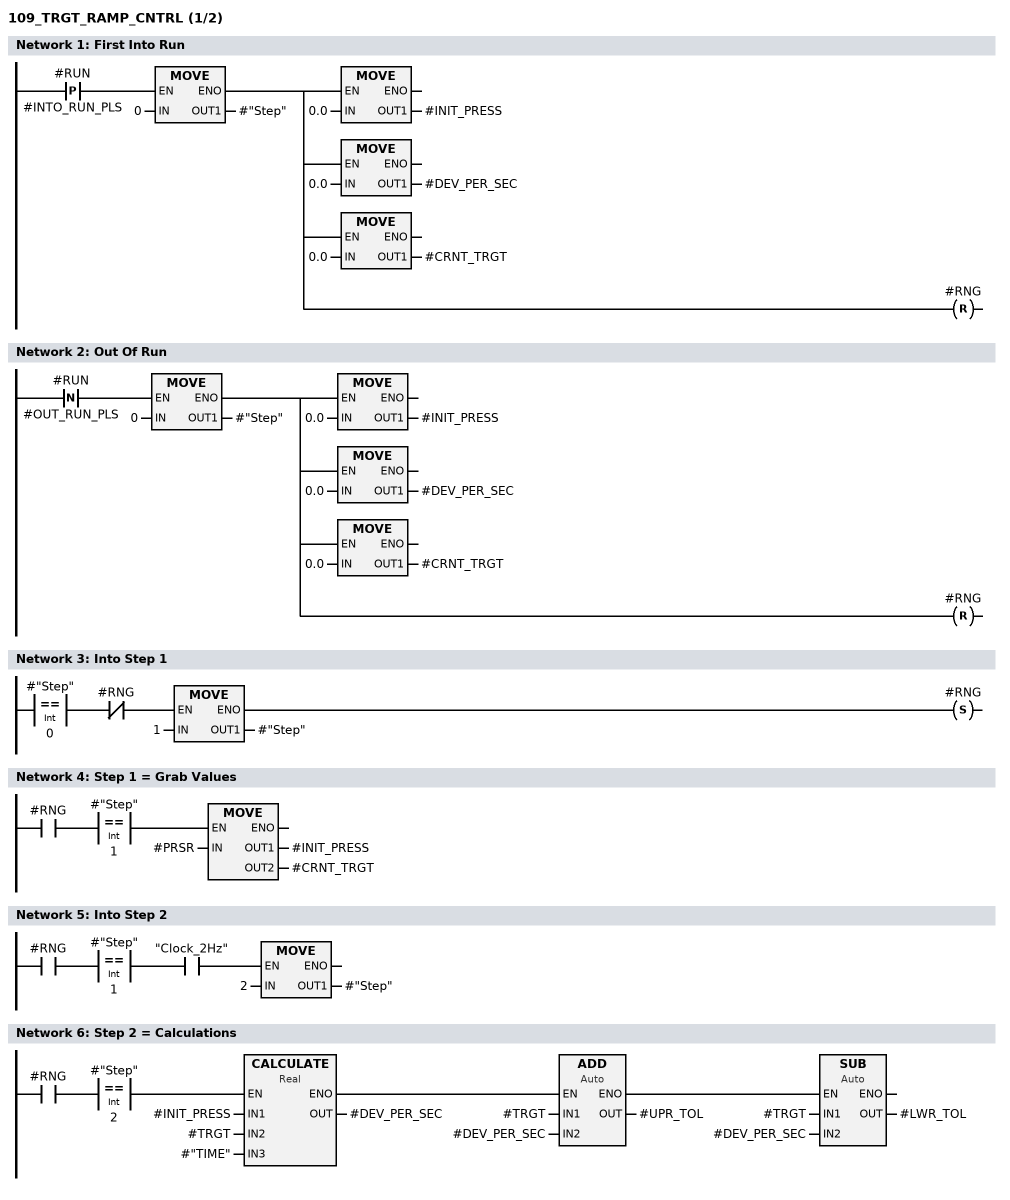
   RUNG wire#powerrail
      P_Contact(operand := #RUN, bit := #INTO_RUN_PLS)
      Move(in := 0, out1 => #"Step")
      wire#w1
      Move(in := 0.0, out1 => #INIT_PRESS)
   END_RUNG
   RUNG wire#w1
      Move(in := 0.0, out1 => #DEV_PER_SEC)
   END_RUNG
   RUNG wire#w1
      Move(in := 0.0, out1 => #CRNT_TRGT)
   END_RUNG
   RUNG wire#w1
      R_Coil( #RNG )
   END_RUNG
   // the same network as SCL:
   #_w1 := #RUN AND NOT #INTO_RUN_PLS;   // rising edge of #RUN
   #INTO_RUN_PLS := #RUN;
   IF #_w1 THEN
       #"Step" := 0;
       #INIT_PRESS := 0.0;
       #DEV_PER_SEC := 0.0;
       #CRNT_TRGT := 0.0;
       #RNG := FALSE;
   END_IF;
END_REGION

REGION Network 2: Out Of Run
   RUNG wire#powerrail
      N_Contact(operand := #RUN, bit := #OUT_RUN_PLS)
      Move(in := 0, out1 => #"Step")
      wire#w1
      Move(in := 0.0, out1 => #INIT_PRESS)
   END_RUNG
   RUNG wire#w1
      Move(in := 0.0, out1 => #DEV_PER_SEC)
   END_RUNG
   RUNG wire#w1
      Move(in := 0.0, out1 => #CRNT_TRGT)
   END_RUNG
   RUNG wire#w1
      R_Coil( #RNG )
   END_RUNG
   // the same network as SCL:
   #_w1 := NOT #RUN AND #OUT_RUN_PLS;   // falling edge of #RUN
   #OUT_RUN_PLS := #RUN;
   IF #_w1 THEN
       #"Step" := 0;
       #INIT_PRESS := 0.0;
       #DEV_PER_SEC := 0.0;
       #CRNT_TRGT := 0.0;
       #RNG := FALSE;
   END_IF;
END_REGION

REGION Network 3: Into Step 1
   RUNG wire#powerrail
      { S7_Templates := "SrcType := Int" } EQ_Contact(in1 := #"Step", in2 := 0)
      I_Contact( #RNG )
      Move(in := 1, out1 => #"Step")
      S_Coil( #RNG )
   END_RUNG
   // the same network as SCL:
   #_w1 := (#"Step" = 0) AND NOT #RNG;
   IF #_w1 THEN
       #"Step" := 1;
       #RNG := TRUE;
   END_IF;
END_REGION

REGION Network 4: Step 1 = Grab Values
   RUNG wire#powerrail
      Contact( #RNG )
      { S7_Templates := "SrcType := Int" } EQ_Contact(in1 := #"Step", in2 := 1)
      Move(in := #PRSR, out1 => #INIT_PRESS, out2 => #CRNT_TRGT)
   END_RUNG
   // the same network as SCL:
   IF #RNG AND (#"Step" = 1) THEN
       #INIT_PRESS := #PRSR;
       #CRNT_TRGT := #PRSR;
   END_IF;
END_REGION

REGION Network 5: Into Step 2
   RUNG wire#powerrail
      Contact( #RNG )
      { S7_Templates := "SrcType := Int" } EQ_Contact(in1 := #"Step", in2 := 1)
      Contact( "Clock_2Hz" )
      Move(in := 2, out1 => #"Step")
   END_RUNG
   // the same network as SCL:
   IF #RNG AND (#"Step" = 1) AND "Clock_2Hz" THEN #"Step" := 2; END_IF;
END_REGION

REGION Network 6: Step 2 = Calculations
   RUNG wire#powerrail
      Contact( #RNG )
      { S7_Templates := "SrcType := Int" } EQ_Contact(in1 := #"Step", in2 := 2)
      { S7_Templates := "SrcType := Real"; S7_Expression := "(IN2-IN1)/IN3" } Calculate(in1 := #INIT_PRESS, in2 := #TRGT, in3 := #"TIME", out => #DEV_PER_SEC)
      Add(in1 := #TRGT, in2 := #DEV_PER_SEC, out => #UPR_TOL)
      Sub(in1 := #TRGT, in2 := #DEV_PER_SEC, out => #LWR_TOL)
   END_RUNG
   // the same network as SCL:
   IF #RNG AND (#"Step" = 2) THEN
       #DEV_PER_SEC := (#TRGT-#INIT_PRESS)/#"TIME";
       #UPR_TOL := #TRGT + #DEV_PER_SEC;
       #LWR_TOL := #TRGT - #DEV_PER_SEC;
   END_IF;
END_REGION

REGION Network 7: Into Step 3 If Ramp Up Needed, Step 4 If Ramp Down Needed, Else Step 5
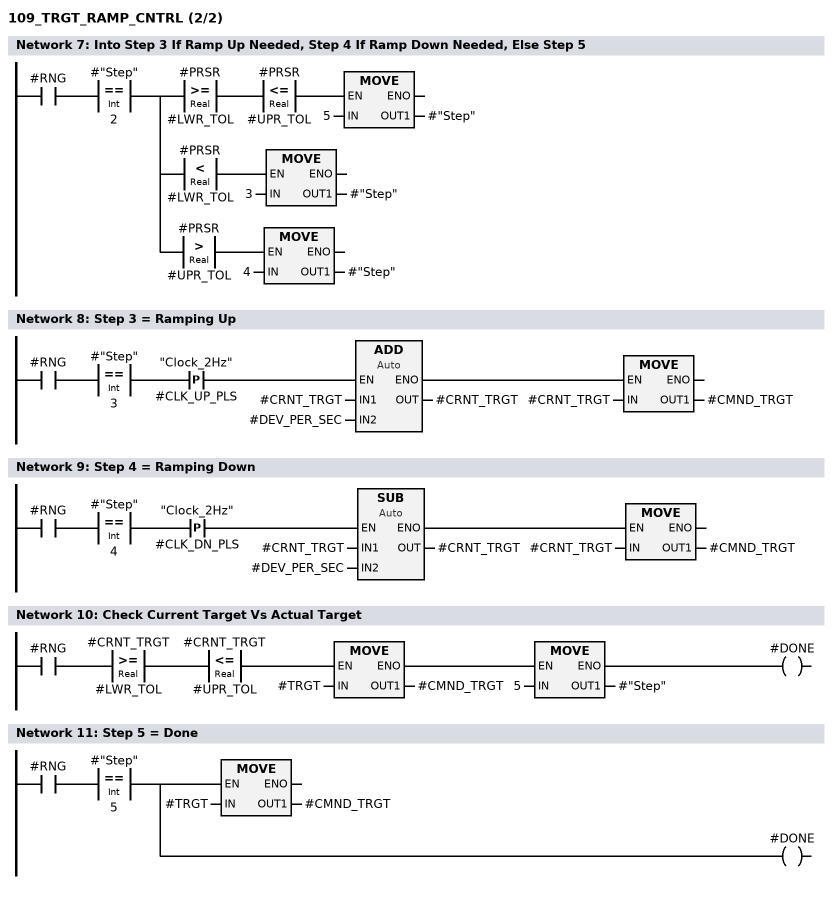
   RUNG wire#powerrail
      Contact( #RNG )
      { S7_Templates := "SrcType := Int" } EQ_Contact(in1 := #"Step", in2 := 2)
      wire#w1
      { S7_Templates := "SrcType := Real" } GE_Contact(in1 := #PRSR, in2 := #LWR_TOL)
      { S7_Templates := "SrcType := Real" } LE_Contact(in1 := #PRSR, in2 := #UPR_TOL)
      Move(in := 5, out1 => #"Step")
   END_RUNG
   RUNG wire#w1
      { S7_Templates := "SrcType := Real" } LT_Contact(in1 := #PRSR, in2 := #LWR_TOL)
      Move(in := 3, out1 => #"Step")
   END_RUNG
   RUNG wire#w1
      { S7_Templates := "SrcType := Real" } GT_Contact(in1 := #PRSR, in2 := #UPR_TOL)
      Move(in := 4, out1 => #"Step")
   END_RUNG
   // the same network as SCL:
   #_w1 := #RNG AND (#"Step" = 2);
   IF #_w1 AND (#PRSR >= #LWR_TOL) AND (#PRSR <= #UPR_TOL) THEN #"Step" := 5; END_IF;
   IF #_w1 AND (#PRSR < #LWR_TOL) THEN #"Step" := 3; END_IF;
   IF #_w1 AND (#PRSR > #UPR_TOL) THEN #"Step" := 4; END_IF;
END_REGION

REGION Network 8: Step 3 = Ramping Up
   RUNG wire#powerrail
      Contact( #RNG )
      { S7_Templates := "SrcType := Int" } EQ_Contact(in1 := #"Step", in2 := 3)
      P_Contact(operand := "Clock_2Hz", bit := #CLK_UP_PLS)
      Add(in1 := #CRNT_TRGT, in2 := #DEV_PER_SEC, out => #CRNT_TRGT)
      Move(in := #CRNT_TRGT, out1 => #CMND_TRGT)
   END_RUNG
   // the same network as SCL:
   #_w1 := #RNG AND (#"Step" = 3) AND "Clock_2Hz" AND NOT #CLK_UP_PLS;   // rising edge of "Clock_2Hz"
   #CLK_UP_PLS := "Clock_2Hz";
   IF #_w1 THEN
       #CRNT_TRGT := #CRNT_TRGT + #DEV_PER_SEC;
       #CMND_TRGT := #CRNT_TRGT;
   END_IF;
END_REGION

REGION Network 9: Step 4 = Ramping Down
   RUNG wire#powerrail
      Contact( #RNG )
      { S7_Templates := "SrcType := Int" } EQ_Contact(in1 := #"Step", in2 := 4)
      P_Contact(operand := "Clock_2Hz", bit := #CLK_DN_PLS)
      Sub(in1 := #CRNT_TRGT, in2 := #DEV_PER_SEC, out => #CRNT_TRGT)
      Move(in := #CRNT_TRGT, out1 => #CMND_TRGT)
   END_RUNG
   // the same network as SCL:
   #_w1 := #RNG AND (#"Step" = 4) AND "Clock_2Hz" AND NOT #CLK_DN_PLS;   // rising edge of "Clock_2Hz"
   #CLK_DN_PLS := "Clock_2Hz";
   IF #_w1 THEN
       #CRNT_TRGT := #CRNT_TRGT - #DEV_PER_SEC;
       #CMND_TRGT := #CRNT_TRGT;
   END_IF;
END_REGION

REGION Network 10: Check Current Target Vs Actual Target
   RUNG wire#powerrail
      Contact( #RNG )
      { S7_Templates := "SrcType := Real" } GE_Contact(in1 := #CRNT_TRGT, in2 := #LWR_TOL)
      { S7_Templates := "SrcType := Real" } LE_Contact(in1 := #CRNT_TRGT, in2 := #UPR_TOL)
      Move(in := #TRGT, out1 => #CMND_TRGT)
      Move(in := 5, out1 => #"Step")
      Coil( #DONE )
   END_RUNG
   // the same network as SCL:
   #_w1 := #RNG AND (#CRNT_TRGT >= #LWR_TOL) AND (#CRNT_TRGT <= #UPR_TOL);
   IF #_w1 THEN
       #CMND_TRGT := #TRGT;
       #"Step" := 5;
   END_IF;
   #DONE := #_w1;
END_REGION

REGION Network 11: Step 5 = Done
   RUNG wire#powerrail
      Contact( #RNG )
      { S7_Templates := "SrcType := Int" } EQ_Contact(in1 := #"Step", in2 := 5)
      wire#w1
      Move(in := #TRGT, out1 => #CMND_TRGT)
   END_RUNG
   RUNG wire#w1
      Coil( #DONE )
   END_RUNG
   // the same network as SCL:
   #_w1 := #RNG AND (#"Step" = 5);
   IF #_w1 THEN #CMND_TRGT := #TRGT; END_IF;
   #DONE := #_w1;
END_REGION
END_FUNCTION_BLOCK

FUNCTION_BLOCK "110_GCU_TNK_FLUSH_SEQ"   // FB110, LAD
TITLE = GCU Tank Flush Sequence
{ S7_Optimized_Access := 'TRUE' }
AUTHOR : JRS
VERSION : 0.1
// For the automatic flushing of the GCU tank
   VAR_INPUT
      RUN : Bool;   // Block control
      FLUSH_TIME : Time := T#60s;   // Flush time
      P305_PRSNT : Bool;   // P305 Fitted
      P305_RNG : Bool;   // Pump running
      P304_RNG : Bool;   // Pump running
      CV358_OPN : Bool;   // Valve open
      CV358_CLSD : Bool;   // Valve closed
   END_VAR
   VAR_OUTPUT
      RUN_P305 : Bool;   // Pump control
      RUN_P304 : Bool;   // Pump control
      OPEN_CV358 : Bool;   // Valve control
      FLUSHING : Bool;   // Flushing status
      DONE : Bool;   // Flushing complete
   END_VAR
   VAR
      INTO_RUN_PLS : Bool;   // Pulse bit
      "STEP" : Int;   // Step number
      RNG : Bool;   // Running bit
      OUT_RUN_PLS : Bool;   // Pulse bit
      CV358_OPND_PAUSE : TON_TIME;   // Pause timer
      P305_RNG_PAUSE : TON_TIME;   // Pause timer
      P304_RNG_PAUSE : TON_TIME;   // Pause timer
      P305_STPD_PAUSE : TON_TIME;   // Pause timer
      P304_STPD_PAUSE : TON_TIME;   // Pause timer
      CV358_CLSD_PAUSE : TON_TIME;   // Pause timer
      FLUSH_TIMER : TON_TIME;   // Flushing time
      "P304_RNG_PAUSE II" : TON_TIME;
   END_VAR
   VAR_TEMP   // added for the SCL form of the ladder/FBD networks
      _w1 : Bool;
   END_VAR
   // CV358_OPND_PAUSE.PT := T#5s;
   // P305_RNG_PAUSE.PT := T#5s;
   // P304_RNG_PAUSE.PT := T#5s;
   // P305_STPD_PAUSE.PT := T#5s;
   // P304_STPD_PAUSE.PT := T#5s;
   // CV358_CLSD_PAUSE.PT := T#5s;
BEGIN

REGION Network 1: First Into Run
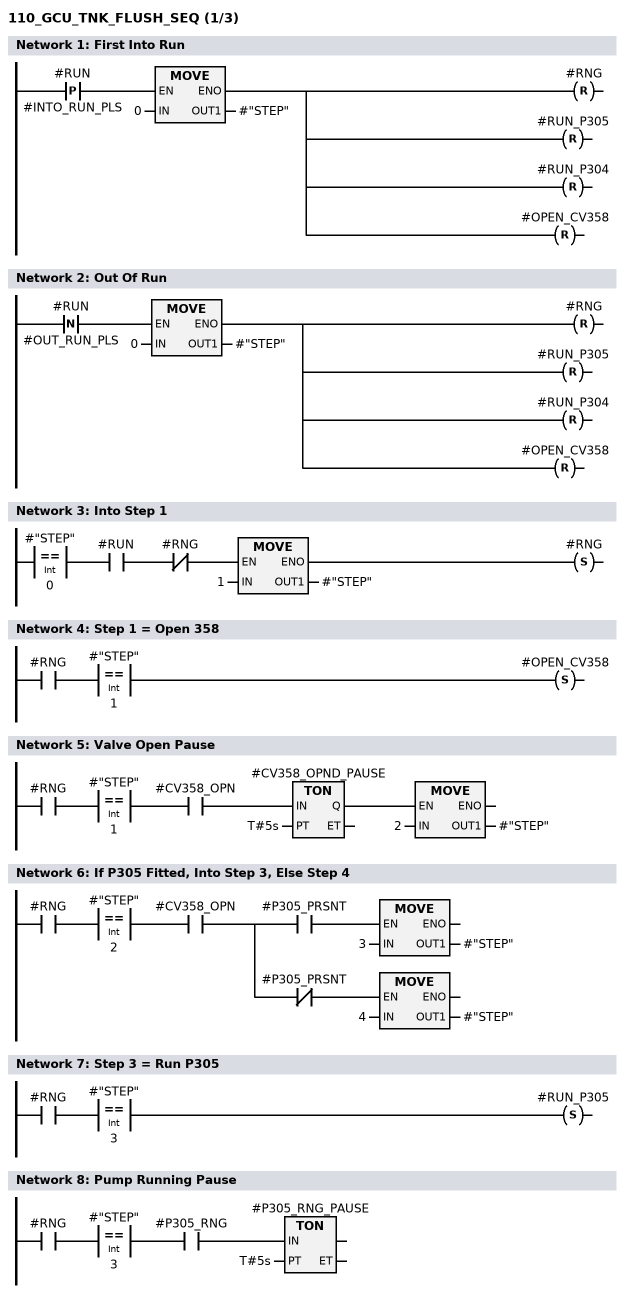
   RUNG wire#powerrail
      P_Contact(operand := #RUN, bit := #INTO_RUN_PLS)
      Move(in := 0, out1 => #"STEP")
      wire#w1
      R_Coil( #RNG )
   END_RUNG
   RUNG wire#w1
      R_Coil( #RUN_P305 )
   END_RUNG
   RUNG wire#w1
      R_Coil( #RUN_P304 )
   END_RUNG
   RUNG wire#w1
      R_Coil( #OPEN_CV358 )
   END_RUNG
   // the same network as SCL:
   #_w1 := #RUN AND NOT #INTO_RUN_PLS;   // rising edge of #RUN
   #INTO_RUN_PLS := #RUN;
   IF #_w1 THEN
       #"STEP" := 0;
       #RNG := FALSE;
       #RUN_P305 := FALSE;
       #RUN_P304 := FALSE;
       #OPEN_CV358 := FALSE;
   END_IF;
END_REGION

REGION Network 2: Out Of Run
   RUNG wire#powerrail
      N_Contact(operand := #RUN, bit := #OUT_RUN_PLS)
      Move(in := 0, out1 => #"STEP")
      wire#w1
      R_Coil( #RNG )
   END_RUNG
   RUNG wire#w1
      R_Coil( #RUN_P305 )
   END_RUNG
   RUNG wire#w1
      R_Coil( #RUN_P304 )
   END_RUNG
   RUNG wire#w1
      R_Coil( #OPEN_CV358 )
   END_RUNG
   // the same network as SCL:
   #_w1 := NOT #RUN AND #OUT_RUN_PLS;   // falling edge of #RUN
   #OUT_RUN_PLS := #RUN;
   IF #_w1 THEN
       #"STEP" := 0;
       #RNG := FALSE;
       #RUN_P305 := FALSE;
       #RUN_P304 := FALSE;
       #OPEN_CV358 := FALSE;
   END_IF;
END_REGION

REGION Network 3: Into Step 1
   RUNG wire#powerrail
      { S7_Templates := "SrcType := Int" } EQ_Contact(in1 := #"STEP", in2 := 0)
      Contact( #RUN )
      I_Contact( #RNG )
      Move(in := 1, out1 => #"STEP")
      S_Coil( #RNG )
   END_RUNG
   // the same network as SCL:
   #_w1 := (#"STEP" = 0) AND #RUN AND NOT #RNG;
   IF #_w1 THEN
       #"STEP" := 1;
       #RNG := TRUE;
   END_IF;
END_REGION

REGION Network 4: Step 1 = Open 358
   RUNG wire#powerrail
      Contact( #RNG )
      { S7_Templates := "SrcType := Int" } EQ_Contact(in1 := #"STEP", in2 := 1)
      S_Coil( #OPEN_CV358 )
   END_RUNG
   // the same network as SCL:
   IF #RNG AND (#"STEP" = 1) THEN #OPEN_CV358 := TRUE; END_IF;
END_REGION

REGION Network 5: Valve Open Pause
   #CV358_OPND_PAUSE(IN := #RNG AND (#"STEP" = 1) AND #CV358_OPN, PT := T#5s);   // TON
   IF #CV358_OPND_PAUSE.Q THEN #"STEP" := 2; END_IF;
END_REGION

REGION Network 6: If P305 Fitted, Into Step 3, Else Step 4
   RUNG wire#powerrail
      Contact( #RNG )
      { S7_Templates := "SrcType := Int" } EQ_Contact(in1 := #"STEP", in2 := 2)
      Contact( #CV358_OPN )
      wire#w1
      Contact( #P305_PRSNT )
      Move(in := 3, out1 => #"STEP")
   END_RUNG
   RUNG wire#w1
      I_Contact( #P305_PRSNT )
      Move(in := 4, out1 => #"STEP")
   END_RUNG
   // the same network as SCL:
   #_w1 := #RNG AND (#"STEP" = 2) AND #CV358_OPN;
   IF #_w1 AND #P305_PRSNT THEN #"STEP" := 3; END_IF;
   IF #_w1 AND NOT #P305_PRSNT THEN #"STEP" := 4; END_IF;
END_REGION

REGION Network 7: Step 3 = Run P305
   RUNG wire#powerrail
      Contact( #RNG )
      { S7_Templates := "SrcType := Int" } EQ_Contact(in1 := #"STEP", in2 := 3)
      S_Coil( #RUN_P305 )
   END_RUNG
   // the same network as SCL:
   IF #RNG AND (#"STEP" = 3) THEN #RUN_P305 := TRUE; END_IF;
END_REGION

REGION Network 8: Pump Running Pause
   #P305_RNG_PAUSE(IN := #RNG AND (#"STEP" = 3) AND #P305_RNG, PT := T#5s);   // TON
END_REGION

REGION Network 9: Into Step 4
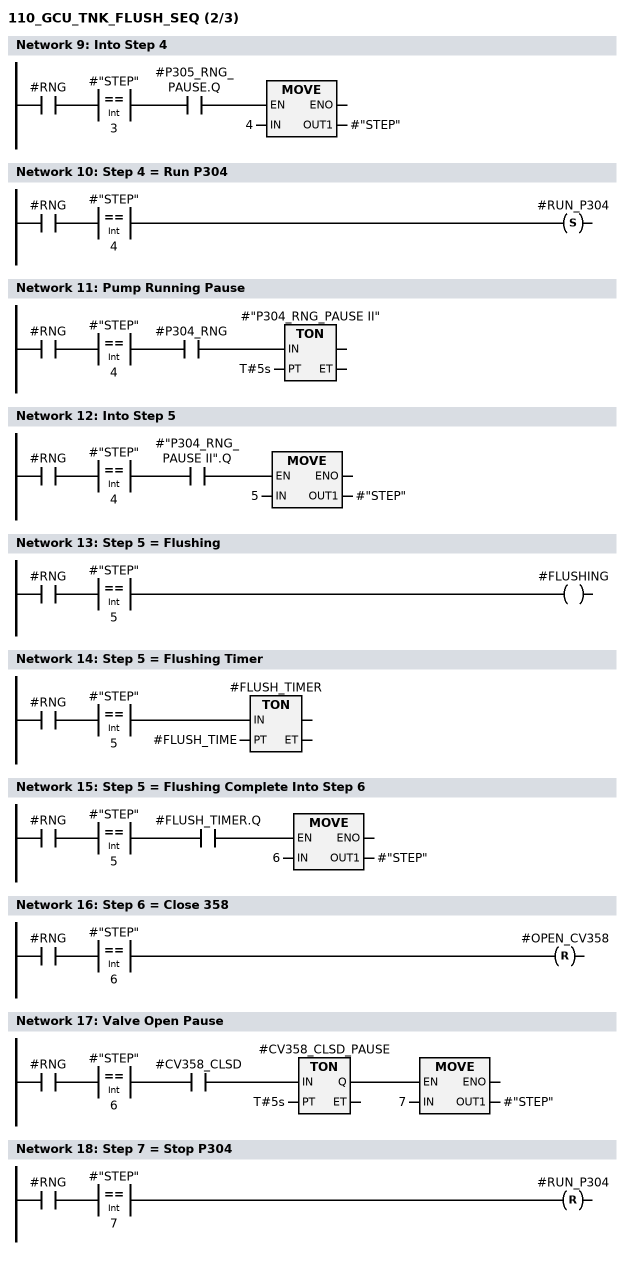
   RUNG wire#powerrail
      Contact( #RNG )
      { S7_Templates := "SrcType := Int" } EQ_Contact(in1 := #"STEP", in2 := 3)
      Contact( #P305_RNG_PAUSE.Q )
      Move(in := 4, out1 => #"STEP")
   END_RUNG
   // the same network as SCL:
   IF #RNG AND (#"STEP" = 3) AND #P305_RNG_PAUSE.Q THEN #"STEP" := 4; END_IF;
END_REGION

REGION Network 10: Step 4 = Run P304
   RUNG wire#powerrail
      Contact( #RNG )
      { S7_Templates := "SrcType := Int" } EQ_Contact(in1 := #"STEP", in2 := 4)
      S_Coil( #RUN_P304 )
   END_RUNG
   // the same network as SCL:
   IF #RNG AND (#"STEP" = 4) THEN #RUN_P304 := TRUE; END_IF;
END_REGION

REGION Network 11: Pump Running Pause
   #"P304_RNG_PAUSE II"(IN := #RNG AND (#"STEP" = 4) AND #P304_RNG, PT := T#5s);   // TON
END_REGION

REGION Network 12: Into Step 5
   RUNG wire#powerrail
      Contact( #RNG )
      { S7_Templates := "SrcType := Int" } EQ_Contact(in1 := #"STEP", in2 := 4)
      Contact( #"P304_RNG_PAUSE II".Q )
      Move(in := 5, out1 => #"STEP")
   END_RUNG
   // the same network as SCL:
   IF #RNG AND (#"STEP" = 4) AND #"P304_RNG_PAUSE II".Q THEN #"STEP" := 5; END_IF;
END_REGION

REGION Network 13: Step 5 = Flushing
   RUNG wire#powerrail
      Contact( #RNG )
      { S7_Templates := "SrcType := Int" } EQ_Contact(in1 := #"STEP", in2 := 5)
      Coil( #FLUSHING )
   END_RUNG
   // the same network as SCL:
   #FLUSHING := #RNG AND (#"STEP" = 5);
END_REGION

REGION Network 14: Step 5 = Flushing Timer
   #FLUSH_TIMER(IN := #RNG AND (#"STEP" = 5), PT := #FLUSH_TIME);   // TON
END_REGION

REGION Network 15: Step 5 = Flushing Complete Into Step 6
   RUNG wire#powerrail
      Contact( #RNG )
      { S7_Templates := "SrcType := Int" } EQ_Contact(in1 := #"STEP", in2 := 5)
      Contact( #FLUSH_TIMER.Q )
      Move(in := 6, out1 => #"STEP")
   END_RUNG
   // the same network as SCL:
   IF #RNG AND (#"STEP" = 5) AND #FLUSH_TIMER.Q THEN #"STEP" := 6; END_IF;
END_REGION

REGION Network 16: Step 6 = Close 358
   RUNG wire#powerrail
      Contact( #RNG )
      { S7_Templates := "SrcType := Int" } EQ_Contact(in1 := #"STEP", in2 := 6)
      R_Coil( #OPEN_CV358 )
   END_RUNG
   // the same network as SCL:
   IF #RNG AND (#"STEP" = 6) THEN #OPEN_CV358 := FALSE; END_IF;
END_REGION

REGION Network 17: Valve Open Pause
   #CV358_CLSD_PAUSE(IN := #RNG AND (#"STEP" = 6) AND #CV358_CLSD, PT := T#5s);   // TON
   IF #CV358_CLSD_PAUSE.Q THEN #"STEP" := 7; END_IF;
END_REGION

REGION Network 18: Step 7 = Stop P304
   RUNG wire#powerrail
      Contact( #RNG )
      { S7_Templates := "SrcType := Int" } EQ_Contact(in1 := #"STEP", in2 := 7)
      R_Coil( #RUN_P304 )
   END_RUNG
   // the same network as SCL:
   IF #RNG AND (#"STEP" = 7) THEN #RUN_P304 := FALSE; END_IF;
END_REGION

REGION Network 19: Pump Stopped Pause
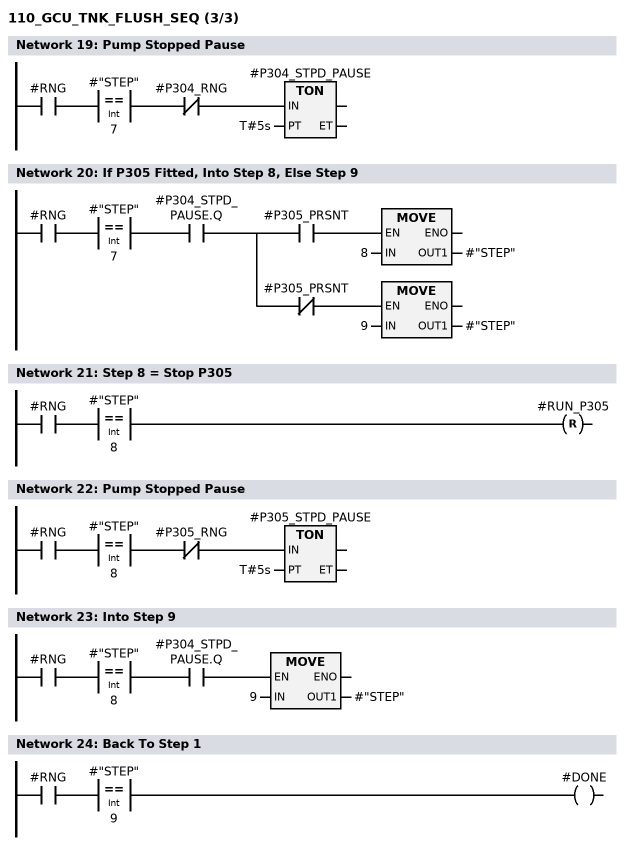
   #P304_STPD_PAUSE(IN := #RNG AND (#"STEP" = 7) AND NOT #P304_RNG, PT := T#5s);   // TON
END_REGION

REGION Network 20: If P305 Fitted, Into Step 8, Else Step 9
   RUNG wire#powerrail
      Contact( #RNG )
      { S7_Templates := "SrcType := Int" } EQ_Contact(in1 := #"STEP", in2 := 7)
      Contact( #P304_STPD_PAUSE.Q )
      wire#w1
      Contact( #P305_PRSNT )
      Move(in := 8, out1 => #"STEP")
   END_RUNG
   RUNG wire#w1
      I_Contact( #P305_PRSNT )
      Move(in := 9, out1 => #"STEP")
   END_RUNG
   // the same network as SCL:
   #_w1 := #RNG AND (#"STEP" = 7) AND #P304_STPD_PAUSE.Q;
   IF #_w1 AND #P305_PRSNT THEN #"STEP" := 8; END_IF;
   IF #_w1 AND NOT #P305_PRSNT THEN #"STEP" := 9; END_IF;
END_REGION

REGION Network 21: Step 8 = Stop P305
   RUNG wire#powerrail
      Contact( #RNG )
      { S7_Templates := "SrcType := Int" } EQ_Contact(in1 := #"STEP", in2 := 8)
      R_Coil( #RUN_P305 )
   END_RUNG
   // the same network as SCL:
   IF #RNG AND (#"STEP" = 8) THEN #RUN_P305 := FALSE; END_IF;
END_REGION

REGION Network 22: Pump Stopped Pause
   #P305_STPD_PAUSE(IN := #RNG AND (#"STEP" = 8) AND NOT #P305_RNG, PT := T#5s);   // TON
END_REGION

REGION Network 23: Into Step 9
   RUNG wire#powerrail
      Contact( #RNG )
      { S7_Templates := "SrcType := Int" } EQ_Contact(in1 := #"STEP", in2 := 8)
      Contact( #P304_STPD_PAUSE.Q )
      Move(in := 9, out1 => #"STEP")
   END_RUNG
   // the same network as SCL:
   IF #RNG AND (#"STEP" = 8) AND #P304_STPD_PAUSE.Q THEN #"STEP" := 9; END_IF;
END_REGION

REGION Network 24: Back To Step 1
   RUNG wire#powerrail
      Contact( #RNG )
      { S7_Templates := "SrcType := Int" } EQ_Contact(in1 := #"STEP", in2 := 9)
      Coil( #DONE )
   END_RUNG
   // the same network as SCL:
   #DONE := #RNG AND (#"STEP" = 9);
END_REGION
END_FUNCTION_BLOCK

FUNCTION_BLOCK "140_PGC_HRS_RUN"   // FB140, LAD
TITLE = PGC Hours Run Control
{ S7_Optimized_Access := 'TRUE' }
AUTHOR : JRS
VERSION : 0.1
// For the recording of hours run and indication of service requirement
   VAR_INPUT
      RUN : Bool;
      RST : Bool;
      SHRS_IP : Int := 1000;
   END_VAR
   VAR_OUTPUT
      HRS : Int;
      MINS : Int;
      SECS : Int;
      SRVC : Bool;
   END_VAR
   VAR_IN_OUT
      SRV_HRS : Int;
   END_VAR
   VAR
      SCND_PLS_1 : Bool;
      SCND_PLS_2 : Bool;
   END_VAR
   VAR RETAIN
      TOT_HRS : Int;
      TOT_MINS : Int;
      TOT_SECS : Int;
      SRV_MIN : Int;
      SRV_SECS : Int;
   END_VAR
   VAR_TEMP   // added for the SCL form of the ladder/FBD networks
      _w1 : Bool;
      _w2 : Bool;
      _w3 : Bool;
   END_VAR
BEGIN

REGION Network 1: Increment Total Hours
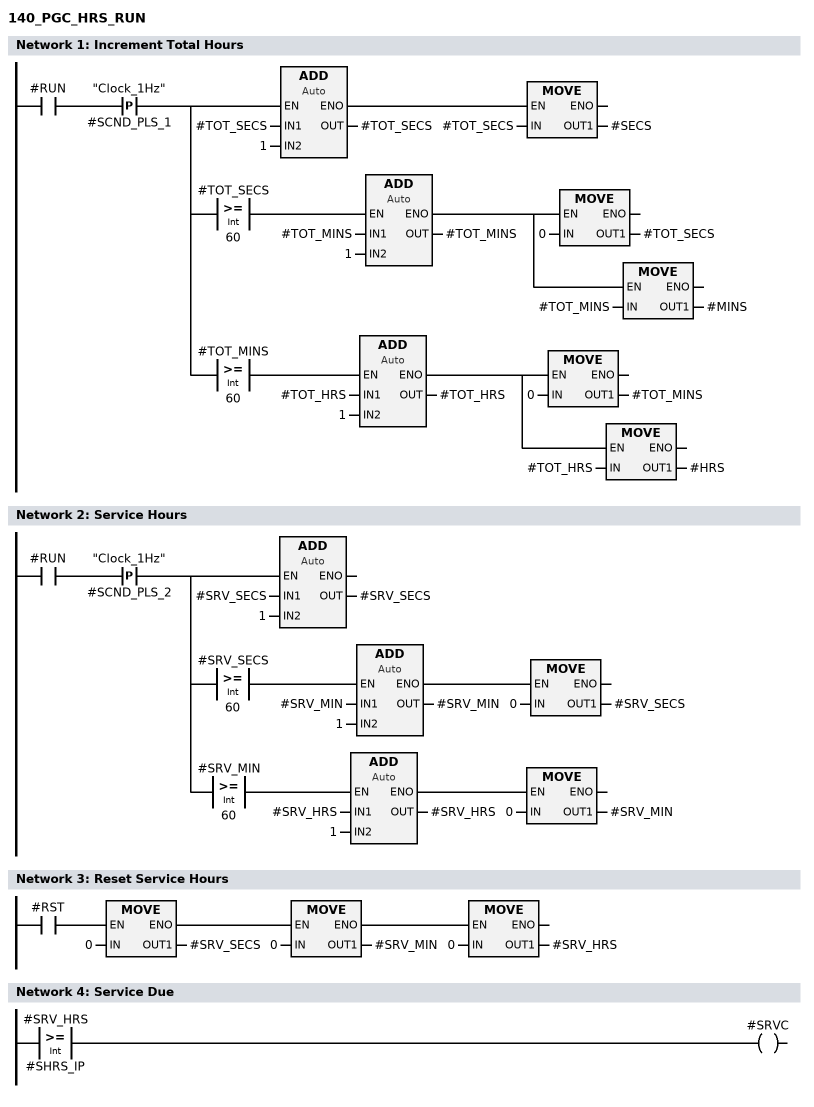
   RUNG wire#powerrail
      Contact( #RUN )
      P_Contact(operand := "Clock_1Hz", bit := #SCND_PLS_1)
      wire#w1
      Add(in1 := #TOT_SECS, in2 := 1, out => #TOT_SECS)
      Move(in := #TOT_SECS, out1 => #SECS)
   END_RUNG
   RUNG wire#w1
      { S7_Templates := "SrcType := Int" } GE_Contact(in1 := #TOT_SECS, in2 := 60)
      Add(in1 := #TOT_MINS, in2 := 1, out => #TOT_MINS)
      wire#w2
      Move(in := 0, out1 => #TOT_SECS)
   END_RUNG
   RUNG wire#w2
      Move(in := #TOT_MINS, out1 => #MINS)
   END_RUNG
   RUNG wire#w1
      { S7_Templates := "SrcType := Int" } GE_Contact(in1 := #TOT_MINS, in2 := 60)
      Add(in1 := #TOT_HRS, in2 := 1, out => #TOT_HRS)
      wire#w3
      Move(in := 0, out1 => #TOT_MINS)
   END_RUNG
   RUNG wire#w3
      Move(in := #TOT_HRS, out1 => #HRS)
   END_RUNG
   // the same network as SCL:
   #_w1 := #RUN AND "Clock_1Hz" AND NOT #SCND_PLS_1;   // rising edge of "Clock_1Hz"
   #SCND_PLS_1 := "Clock_1Hz";
   IF #_w1 THEN
       #TOT_SECS := #TOT_SECS + 1;
       #SECS := #TOT_SECS;
   END_IF;
   IF #_w1 AND (#TOT_SECS >= 60) THEN #TOT_MINS := #TOT_MINS + 1; END_IF;
   #_w2 := #_w1 AND (#TOT_SECS >= 60);
   IF #_w2 THEN
       #TOT_SECS := 0;
       #MINS := #TOT_MINS;
   END_IF;
   IF #_w1 AND (#TOT_MINS >= 60) THEN #TOT_HRS := #TOT_HRS + 1; END_IF;
   #_w3 := #_w1 AND (#TOT_MINS >= 60);
   IF #_w3 THEN
       #TOT_MINS := 0;
       #HRS := #TOT_HRS;
   END_IF;
END_REGION

REGION Network 2: Service Hours
   RUNG wire#powerrail
      Contact( #RUN )
      P_Contact(operand := "Clock_1Hz", bit := #SCND_PLS_2)
      wire#w1
      Add(in1 := #SRV_SECS, in2 := 1, out => #SRV_SECS)
   END_RUNG
   RUNG wire#w1
      { S7_Templates := "SrcType := Int" } GE_Contact(in1 := #SRV_SECS, in2 := 60)
      Add(in1 := #SRV_MIN, in2 := 1, out => #SRV_MIN)
      Move(in := 0, out1 => #SRV_SECS)
   END_RUNG
   RUNG wire#w1
      { S7_Templates := "SrcType := Int" } GE_Contact(in1 := #SRV_MIN, in2 := 60)
      Add(in1 := #SRV_HRS, in2 := 1, out => #SRV_HRS)
      Move(in := 0, out1 => #SRV_MIN)
   END_RUNG
   // the same network as SCL:
   #_w1 := #RUN AND "Clock_1Hz" AND NOT #SCND_PLS_2;   // rising edge of "Clock_1Hz"
   #SCND_PLS_2 := "Clock_1Hz";
   IF #_w1 THEN #SRV_SECS := #SRV_SECS + 1; END_IF;
   IF #_w1 AND (#SRV_SECS >= 60) THEN
       #SRV_MIN := #SRV_MIN + 1;
       #SRV_SECS := 0;
   END_IF;
   IF #_w1 AND (#SRV_MIN >= 60) THEN
       #SRV_HRS := #SRV_HRS + 1;
       #SRV_MIN := 0;
   END_IF;
END_REGION

REGION Network 3: Reset Service Hours
   RUNG wire#powerrail
      Contact( #RST )
      Move(in := 0, out1 => #SRV_SECS)
      Move(in := 0, out1 => #SRV_MIN)
      Move(in := 0, out1 => #SRV_HRS)
   END_RUNG
   // the same network as SCL:
   IF #RST THEN
       #SRV_SECS := 0;
       #SRV_MIN := 0;
       #SRV_HRS := 0;
   END_IF;
END_REGION

REGION Network 4: Service Due
   RUNG wire#powerrail
      { S7_Templates := "SrcType := Int" } GE_Contact(in1 := #SRV_HRS, in2 := #SHRS_IP)
      Coil( #SRVC )
   END_RUNG
   // the same network as SCL:
   #SRVC := #SRV_HRS >= #SHRS_IP;
END_REGION
END_FUNCTION_BLOCK

FUNCTION_BLOCK "141_P303_HRS_RUN"   // FB141, LAD
TITLE = PGC Hours Run Control
{ S7_Optimized_Access := 'TRUE' }
AUTHOR : JRS
VERSION : 0.1
// For the recording of hours run and indication of service requirement
   VAR_INPUT
      RUN : Bool;
      RST : Bool;
      SHRS_IP : Int := 1000;
   END_VAR
   VAR_OUTPUT
      HRS : Int;
      MINS : Int;
      SECS : Int;
      SRVC : Bool;
   END_VAR
   VAR_IN_OUT
      SRV_HRS : Int;
   END_VAR
   VAR
      SCND_PLS_1 : Bool;
      SCND_PLS_2 : Bool;
   END_VAR
   VAR RETAIN
      TOT_HRS : Int;
      TOT_MINS : Int;
      TOT_SECS : Int;
      SRV_MIN : Int;
      SRV_SECS : Int;
   END_VAR
   VAR_TEMP   // added for the SCL form of the ladder/FBD networks
      _w1 : Bool;
      _w2 : Bool;
      _w3 : Bool;
   END_VAR
BEGIN

REGION Network 1: Increment Total Hours
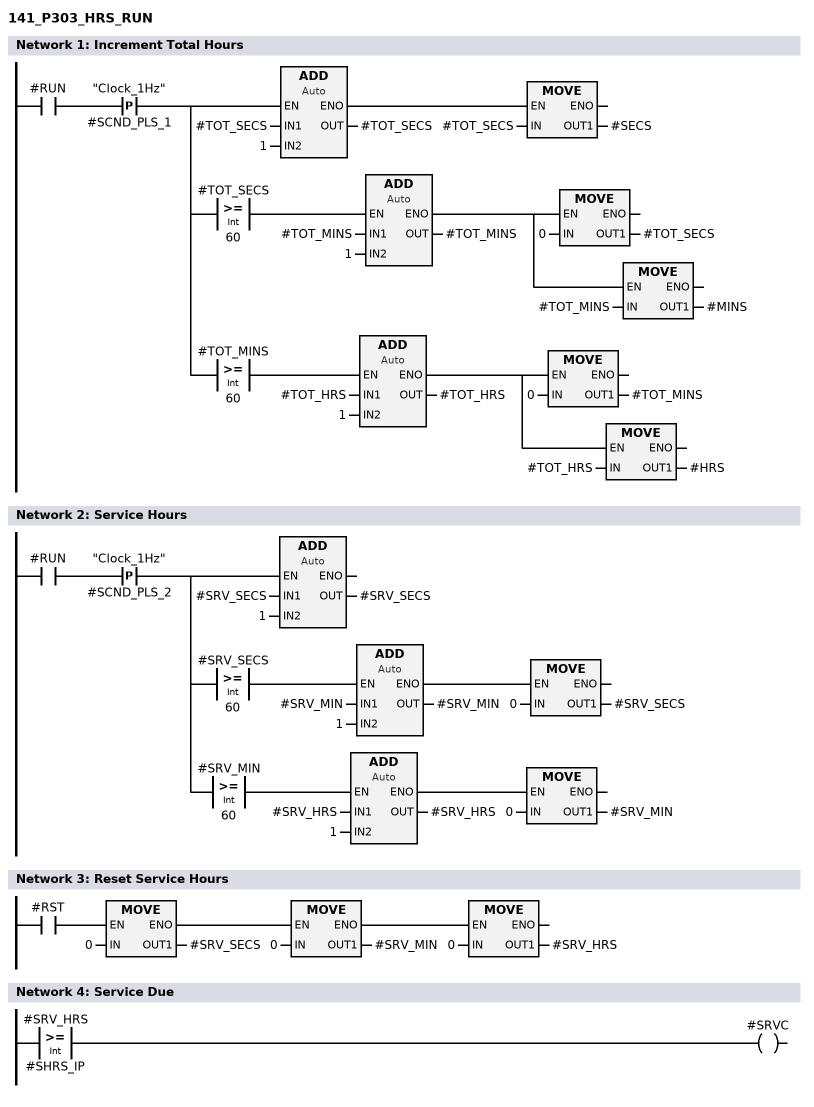
   RUNG wire#powerrail
      Contact( #RUN )
      P_Contact(operand := "Clock_1Hz", bit := #SCND_PLS_1)
      wire#w1
      Add(in1 := #TOT_SECS, in2 := 1, out => #TOT_SECS)
      Move(in := #TOT_SECS, out1 => #SECS)
   END_RUNG
   RUNG wire#w1
      { S7_Templates := "SrcType := Int" } GE_Contact(in1 := #TOT_SECS, in2 := 60)
      Add(in1 := #TOT_MINS, in2 := 1, out => #TOT_MINS)
      wire#w2
      Move(in := 0, out1 => #TOT_SECS)
   END_RUNG
   RUNG wire#w2
      Move(in := #TOT_MINS, out1 => #MINS)
   END_RUNG
   RUNG wire#w1
      { S7_Templates := "SrcType := Int" } GE_Contact(in1 := #TOT_MINS, in2 := 60)
      Add(in1 := #TOT_HRS, in2 := 1, out => #TOT_HRS)
      wire#w3
      Move(in := 0, out1 => #TOT_MINS)
   END_RUNG
   RUNG wire#w3
      Move(in := #TOT_HRS, out1 => #HRS)
   END_RUNG
   // the same network as SCL:
   #_w1 := #RUN AND "Clock_1Hz" AND NOT #SCND_PLS_1;   // rising edge of "Clock_1Hz"
   #SCND_PLS_1 := "Clock_1Hz";
   IF #_w1 THEN
       #TOT_SECS := #TOT_SECS + 1;
       #SECS := #TOT_SECS;
   END_IF;
   IF #_w1 AND (#TOT_SECS >= 60) THEN #TOT_MINS := #TOT_MINS + 1; END_IF;
   #_w2 := #_w1 AND (#TOT_SECS >= 60);
   IF #_w2 THEN
       #TOT_SECS := 0;
       #MINS := #TOT_MINS;
   END_IF;
   IF #_w1 AND (#TOT_MINS >= 60) THEN #TOT_HRS := #TOT_HRS + 1; END_IF;
   #_w3 := #_w1 AND (#TOT_MINS >= 60);
   IF #_w3 THEN
       #TOT_MINS := 0;
       #HRS := #TOT_HRS;
   END_IF;
END_REGION

REGION Network 2: Service Hours
   RUNG wire#powerrail
      Contact( #RUN )
      P_Contact(operand := "Clock_1Hz", bit := #SCND_PLS_2)
      wire#w1
      Add(in1 := #SRV_SECS, in2 := 1, out => #SRV_SECS)
   END_RUNG
   RUNG wire#w1
      { S7_Templates := "SrcType := Int" } GE_Contact(in1 := #SRV_SECS, in2 := 60)
      Add(in1 := #SRV_MIN, in2 := 1, out => #SRV_MIN)
      Move(in := 0, out1 => #SRV_SECS)
   END_RUNG
   RUNG wire#w1
      { S7_Templates := "SrcType := Int" } GE_Contact(in1 := #SRV_MIN, in2 := 60)
      Add(in1 := #SRV_HRS, in2 := 1, out => #SRV_HRS)
      Move(in := 0, out1 => #SRV_MIN)
   END_RUNG
   // the same network as SCL:
   #_w1 := #RUN AND "Clock_1Hz" AND NOT #SCND_PLS_2;   // rising edge of "Clock_1Hz"
   #SCND_PLS_2 := "Clock_1Hz";
   IF #_w1 THEN #SRV_SECS := #SRV_SECS + 1; END_IF;
   IF #_w1 AND (#SRV_SECS >= 60) THEN
       #SRV_MIN := #SRV_MIN + 1;
       #SRV_SECS := 0;
   END_IF;
   IF #_w1 AND (#SRV_MIN >= 60) THEN
       #SRV_HRS := #SRV_HRS + 1;
       #SRV_MIN := 0;
   END_IF;
END_REGION

REGION Network 3: Reset Service Hours
   RUNG wire#powerrail
      Contact( #RST )
      Move(in := 0, out1 => #SRV_SECS)
      Move(in := 0, out1 => #SRV_MIN)
      Move(in := 0, out1 => #SRV_HRS)
   END_RUNG
   // the same network as SCL:
   IF #RST THEN
       #SRV_SECS := 0;
       #SRV_MIN := 0;
       #SRV_HRS := 0;
   END_IF;
END_REGION

REGION Network 4: Service Due
   RUNG wire#powerrail
      { S7_Templates := "SrcType := Int" } GE_Contact(in1 := #SRV_HRS, in2 := #SHRS_IP)
      Coil( #SRVC )
   END_RUNG
   // the same network as SCL:
   #SRVC := #SRV_HRS >= #SHRS_IP;
END_REGION
END_FUNCTION_BLOCK

FUNCTION_BLOCK "142_P304_HRS_RUN"   // FB142, LAD
TITLE = PGC Hours Run Control
{ S7_Optimized_Access := 'TRUE' }
AUTHOR : JRS
VERSION : 0.1
// For the recording of hours run and indication of service requirement
   VAR_INPUT
      RUN : Bool;
      RST : Bool;
      SHRS_IP : Int := 1000;
   END_VAR
   VAR_OUTPUT
      HRS : Int;
      MINS : Int;
      SECS : Int;
      SRVC : Bool;
   END_VAR
   VAR_IN_OUT
      SRV_HRS : Int;
   END_VAR
   VAR
      SCND_PLS_1 : Bool;
      SCND_PLS_2 : Bool;
   END_VAR
   VAR RETAIN
      TOT_HRS : Int;
      TOT_MINS : Int;
      TOT_SECS : Int;
      SRV_MIN : Int;
      SRV_SECS : Int;
   END_VAR
   VAR_TEMP   // added for the SCL form of the ladder/FBD networks
      _w1 : Bool;
      _w2 : Bool;
      _w3 : Bool;
   END_VAR
BEGIN

REGION Network 1: Increment Total Hours
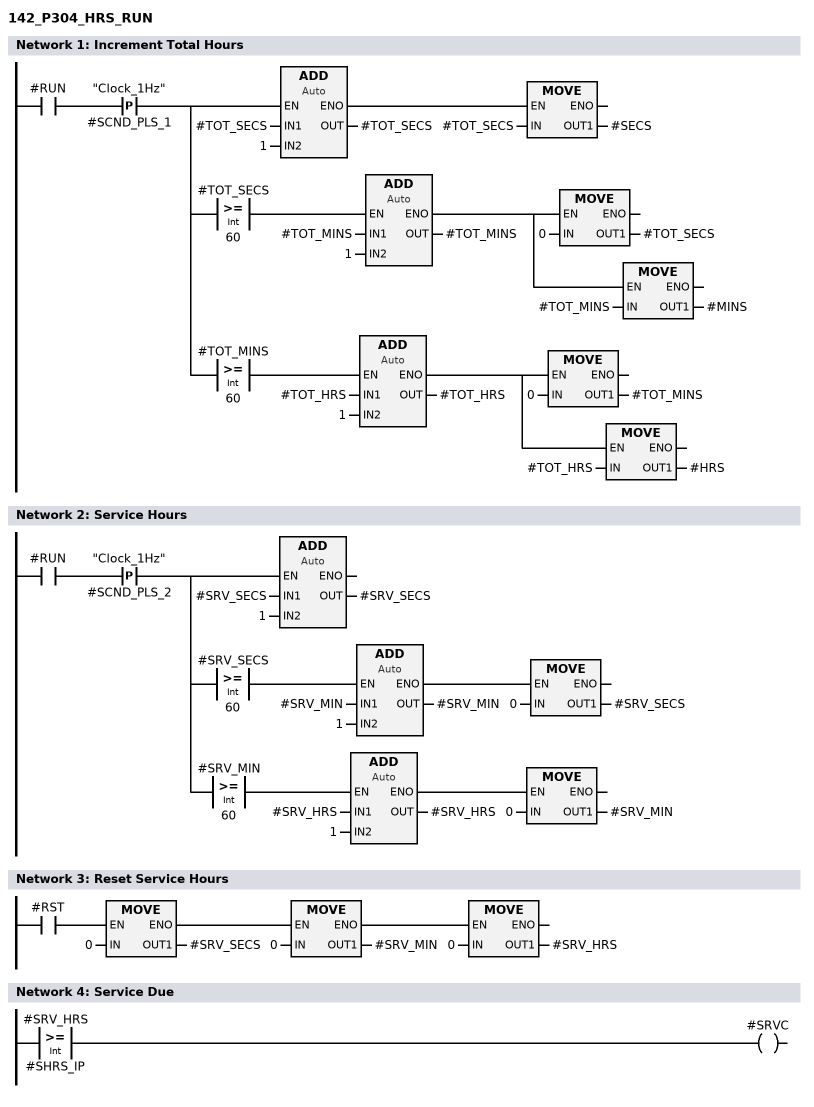
   RUNG wire#powerrail
      Contact( #RUN )
      P_Contact(operand := "Clock_1Hz", bit := #SCND_PLS_1)
      wire#w1
      Add(in1 := #TOT_SECS, in2 := 1, out => #TOT_SECS)
      Move(in := #TOT_SECS, out1 => #SECS)
   END_RUNG
   RUNG wire#w1
      { S7_Templates := "SrcType := Int" } GE_Contact(in1 := #TOT_SECS, in2 := 60)
      Add(in1 := #TOT_MINS, in2 := 1, out => #TOT_MINS)
      wire#w2
      Move(in := 0, out1 => #TOT_SECS)
   END_RUNG
   RUNG wire#w2
      Move(in := #TOT_MINS, out1 => #MINS)
   END_RUNG
   RUNG wire#w1
      { S7_Templates := "SrcType := Int" } GE_Contact(in1 := #TOT_MINS, in2 := 60)
      Add(in1 := #TOT_HRS, in2 := 1, out => #TOT_HRS)
      wire#w3
      Move(in := 0, out1 => #TOT_MINS)
   END_RUNG
   RUNG wire#w3
      Move(in := #TOT_HRS, out1 => #HRS)
   END_RUNG
   // the same network as SCL:
   #_w1 := #RUN AND "Clock_1Hz" AND NOT #SCND_PLS_1;   // rising edge of "Clock_1Hz"
   #SCND_PLS_1 := "Clock_1Hz";
   IF #_w1 THEN
       #TOT_SECS := #TOT_SECS + 1;
       #SECS := #TOT_SECS;
   END_IF;
   IF #_w1 AND (#TOT_SECS >= 60) THEN #TOT_MINS := #TOT_MINS + 1; END_IF;
   #_w2 := #_w1 AND (#TOT_SECS >= 60);
   IF #_w2 THEN
       #TOT_SECS := 0;
       #MINS := #TOT_MINS;
   END_IF;
   IF #_w1 AND (#TOT_MINS >= 60) THEN #TOT_HRS := #TOT_HRS + 1; END_IF;
   #_w3 := #_w1 AND (#TOT_MINS >= 60);
   IF #_w3 THEN
       #TOT_MINS := 0;
       #HRS := #TOT_HRS;
   END_IF;
END_REGION

REGION Network 2: Service Hours
   RUNG wire#powerrail
      Contact( #RUN )
      P_Contact(operand := "Clock_1Hz", bit := #SCND_PLS_2)
      wire#w1
      Add(in1 := #SRV_SECS, in2 := 1, out => #SRV_SECS)
   END_RUNG
   RUNG wire#w1
      { S7_Templates := "SrcType := Int" } GE_Contact(in1 := #SRV_SECS, in2 := 60)
      Add(in1 := #SRV_MIN, in2 := 1, out => #SRV_MIN)
      Move(in := 0, out1 => #SRV_SECS)
   END_RUNG
   RUNG wire#w1
      { S7_Templates := "SrcType := Int" } GE_Contact(in1 := #SRV_MIN, in2 := 60)
      Add(in1 := #SRV_HRS, in2 := 1, out => #SRV_HRS)
      Move(in := 0, out1 => #SRV_MIN)
   END_RUNG
   // the same network as SCL:
   #_w1 := #RUN AND "Clock_1Hz" AND NOT #SCND_PLS_2;   // rising edge of "Clock_1Hz"
   #SCND_PLS_2 := "Clock_1Hz";
   IF #_w1 THEN #SRV_SECS := #SRV_SECS + 1; END_IF;
   IF #_w1 AND (#SRV_SECS >= 60) THEN
       #SRV_MIN := #SRV_MIN + 1;
       #SRV_SECS := 0;
   END_IF;
   IF #_w1 AND (#SRV_MIN >= 60) THEN
       #SRV_HRS := #SRV_HRS + 1;
       #SRV_MIN := 0;
   END_IF;
END_REGION

REGION Network 3: Reset Service Hours
   RUNG wire#powerrail
      Contact( #RST )
      Move(in := 0, out1 => #SRV_SECS)
      Move(in := 0, out1 => #SRV_MIN)
      Move(in := 0, out1 => #SRV_HRS)
   END_RUNG
   // the same network as SCL:
   IF #RST THEN
       #SRV_SECS := 0;
       #SRV_MIN := 0;
       #SRV_HRS := 0;
   END_IF;
END_REGION

REGION Network 4: Service Due
   RUNG wire#powerrail
      { S7_Templates := "SrcType := Int" } GE_Contact(in1 := #SRV_HRS, in2 := #SHRS_IP)
      Coil( #SRVC )
   END_RUNG
   // the same network as SCL:
   #SRVC := #SRV_HRS >= #SHRS_IP;
END_REGION
END_FUNCTION_BLOCK

FUNCTION "100_SC" : Void   // FC100, LAD
TITLE = State Complete
{ S7_Optimized_Access := 'TRUE' }
AUTHOR : JRS
VERSION : 0.1
// For the determination of each step state being complete
   VAR_TEMP   // added for the SCL form of the ladder/FBD networks
      _w1 : Bool;
   END_VAR
BEGIN

REGION Network 1: Step 001 = Confirm Auto Conditions Ok